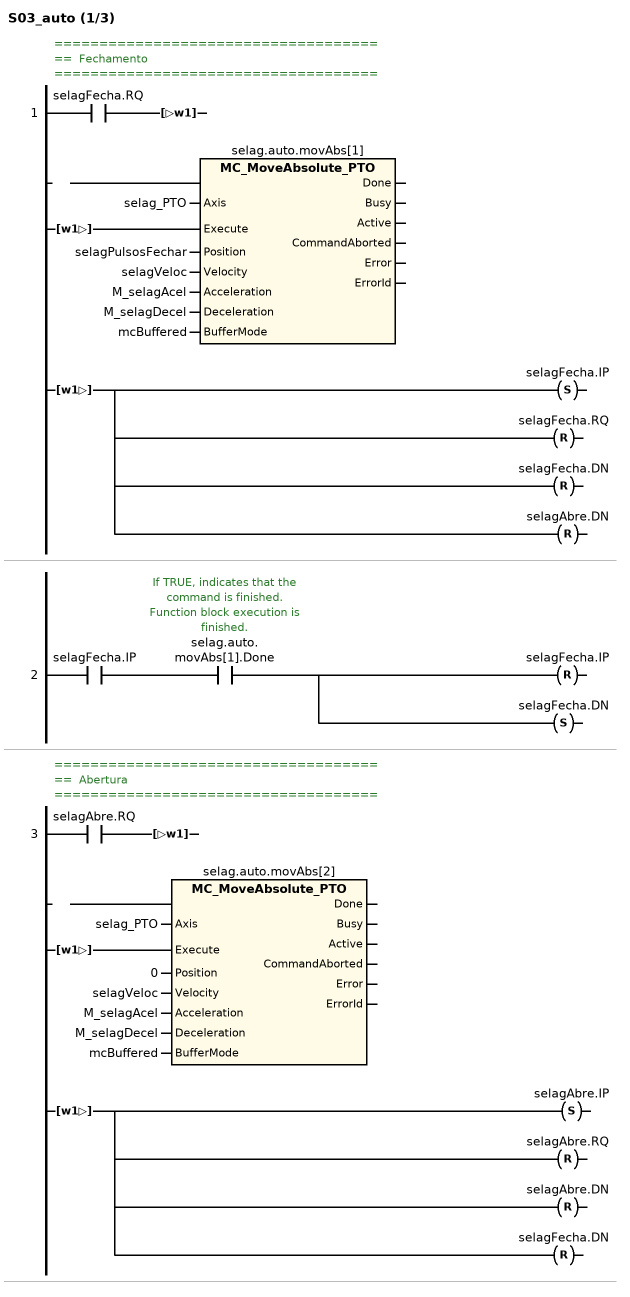
// NETWORK 1
// ====================================
// ==  Fechamento
// ====================================
_w1 := selagFecha.RQ;
selag.auto.movAbs[1](
    Axis := selag_PTO,
    Execute := _w1,
    Position := selagPulsosFechar,
    Velocity := selagVeloc,
    Acceleration := M_selagAcel,
    Deceleration := M_selagDecel,
    BufferMode := mcBuffered); // MC_MoveAbsolute_PTO
selagFecha.IP S= _w1;
selagFecha.RQ R= _w1;
selagFecha.DN R= _w1;
selagAbre.DN R= _w1;

// NETWORK 2
//   selag.auto.movAbs[1].Done: If TRUE, indicates that the command is finished. Function block execution is finished.
_w2 := selagFecha.IP AND selag.auto.movAbs[1].Done;
selagFecha.IP R= _w2;
selagFecha.DN S= _w2;

// NETWORK 3
// ====================================
// ==  Abertura
// ====================================
_w3 := selagAbre.RQ;
selag.auto.movAbs[2](
    Axis := selag_PTO,
    Execute := _w3,
    Position := 0,
    Velocity := selagVeloc,
    Acceleration := M_selagAcel,
    Deceleration := M_selagDecel,
    BufferMode := mcBuffered); // MC_MoveAbsolute_PTO
selagAbre.IP S= _w3;
selagAbre.RQ R= _w3;
selagAbre.DN R= _w3;
selagFecha.DN R= _w3;

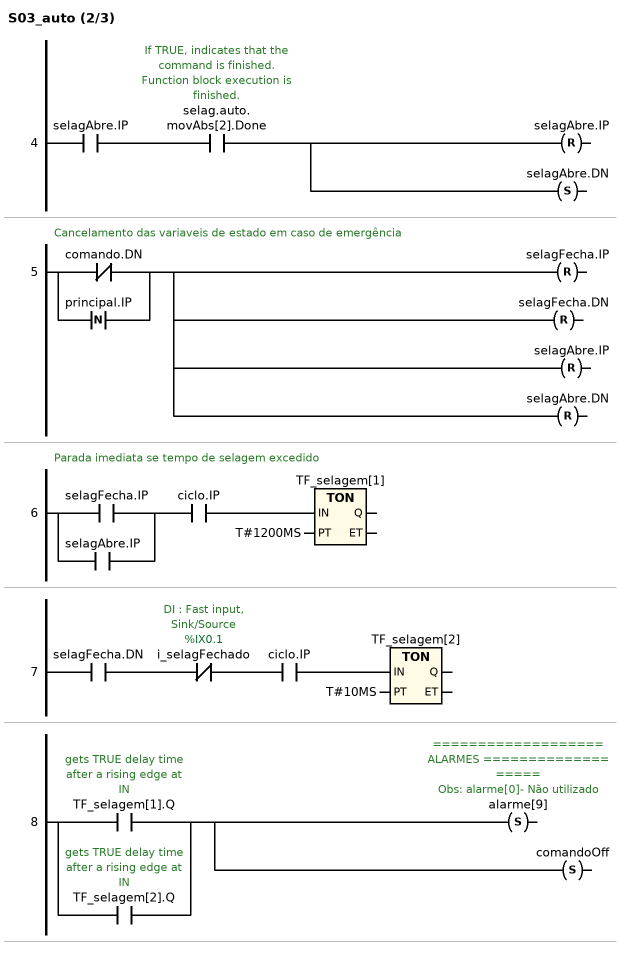
// NETWORK 4
//   selag.auto.movAbs[2].Done: If TRUE, indicates that the command is finished. Function block execution is finished.
_w4 := selagAbre.IP AND selag.auto.movAbs[2].Done;
selagAbre.IP R= _w4;
selagAbre.DN S= _w4;

// NETWORK 5
// Cancelamento das variaveis de estado em caso de emergência
_ft1(CLK := principal.IP);
_w5 := NOT comando.DN OR _ft1.Q;
selagFecha.IP R= _w5;
selagFecha.DN R= _w5;
selagAbre.IP R= _w5;
selagAbre.DN R= _w5;

// NETWORK 6
// Parada imediata se tempo de selagem excedido
TF_selagem[1](IN := (selagFecha.IP OR selagAbre.IP) AND ciclo.IP, PT := T#1200MS); // TON

// NETWORK 7
//   i_selagFechado: DI : Fast input, Sink/Source | AT %IX0.1
TF_selagem[2](IN := selagFecha.DN AND NOT i_selagFechado AND ciclo.IP, PT := T#10MS); // TON

// NETWORK 8
//   TF_selagem[1].Q: gets TRUE delay time after a rising edge at IN
//   TF_selagem[2].Q: gets TRUE delay time after a rising edge at IN
//   alarme[9]: =================== ALARMES =================== Obs: alarme[0]- Não utilizado
_w6 := TF_selagem[1].Q OR TF_selagem[2].Q;
alarme[9] S= _w6;
comandoOff S= _w6;

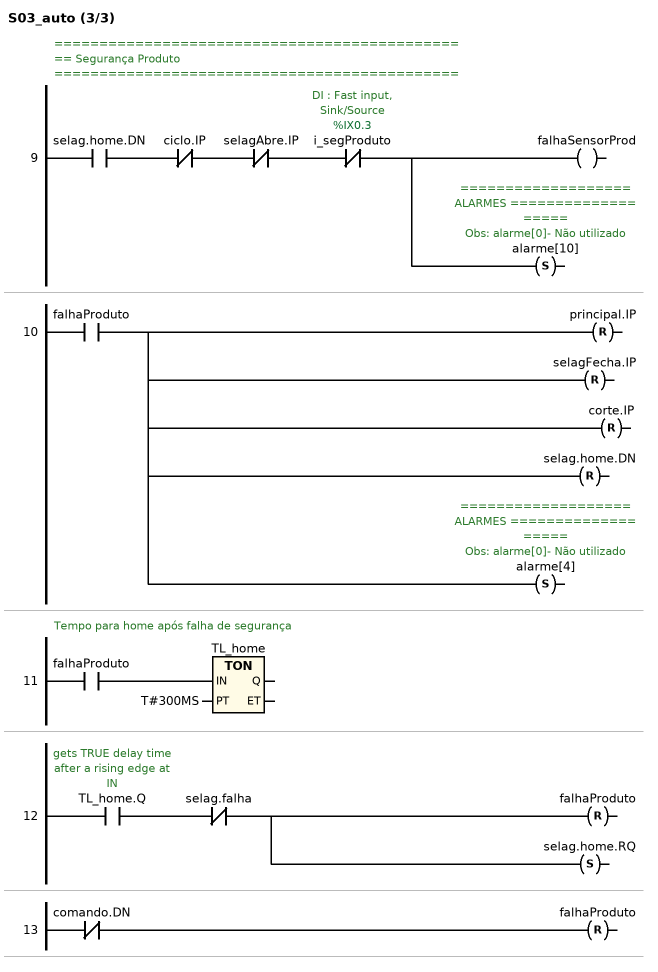
// NETWORK 9
// =============================================
// == Segurança Produto
// =============================================
//   i_segProduto: DI : Fast input, Sink/Source | AT %IX0.3
//   alarme[10]: =================== ALARMES =================== Obs: alarme[0]- Não utilizado
_w7 := selag.home.DN AND NOT ciclo.IP AND NOT selagAbre.IP AND NOT i_segProduto;
falhaSensorProd := _w7;
alarme[10] S= _w7;

// NETWORK 10
//   alarme[4]: =================== ALARMES =================== Obs: alarme[0]- Não utilizado
principal.IP R= falhaProduto;
selagFecha.IP R= falhaProduto;
corte.IP R= falhaProduto;
selag.home.DN R= falhaProduto;
alarme[4] S= falhaProduto;

// NETWORK 11
// Tempo para home após falha de segurança
TL_home(IN := falhaProduto, PT := T#300MS); // TON

// NETWORK 12
//   TL_home.Q: gets TRUE delay time after a rising edge at IN
_w8 := TL_home.Q AND NOT selag.falha;
falhaProduto R= _w8;
selag.home.RQ S= _w8;

// NETWORK 13
falhaProduto R= NOT comando.DN;

END_PROGRAM

// MyController/Application/03_Selagem/S99_calculo
PROGRAM S99_calculo
VAR
END_VAR

selag.calcula:= FALSE;

// cálculo do num pulsos/mm - 1volta motor = 47 mm
selagPulsosMm:= M_selagPulsosVolta / 47;

// cálculo das distâncias a serem percorridas
selagPulsosFechar:= REAL_TO_DINT(M_selagPosFecha * selagPulsosMm / 10);

// cálculo da velocidade
selagVeloc:= 299 * M_selagPulsosVolta * M_selagVeloc / 6000;
selagVelocHome:= 299 * M_selagPulsosVolta * M_selagVelocHome / 6000;

END_PROGRAM

// MyController/Application/04_Disco/D03_auto
PROGRAM D03_auto
VAR
	TF_foto						: TON;
END_VAR
VAR // added by the converter: edge detectors and wires of the graphical bodies
    _w1, _w2 : BOOL;
    _ft1 : F_TRIG;
END_VAR

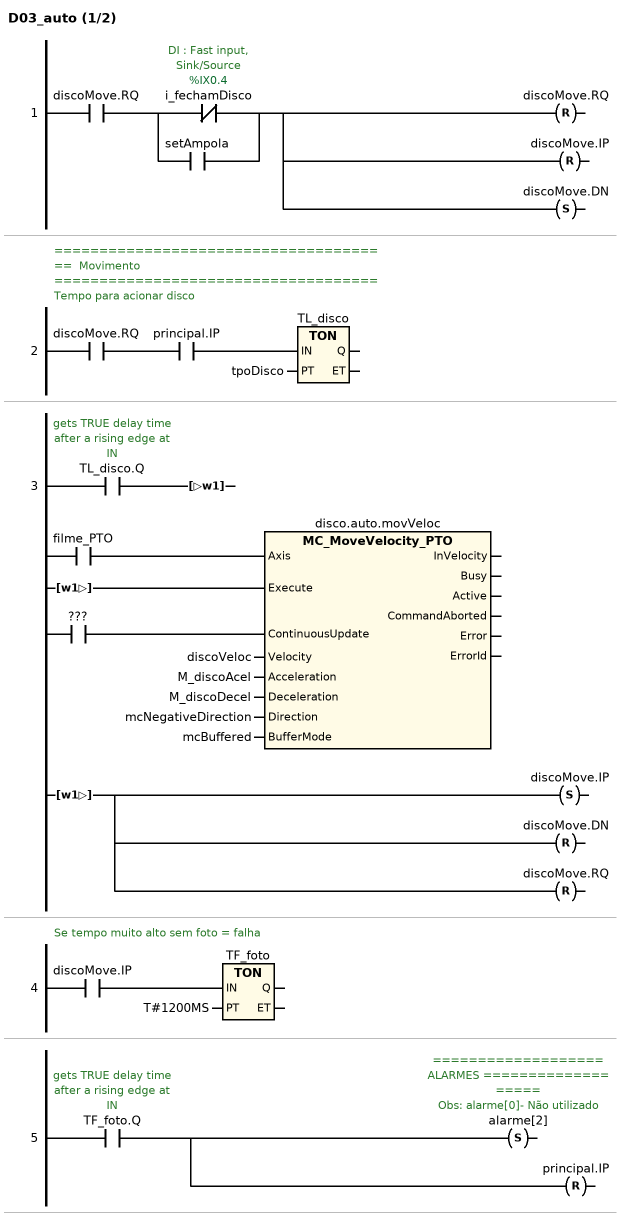
// NETWORK 1
//   i_fechamDisco: DI : Fast input, Sink/Source | AT %IX0.4
_w1 := discoMove.RQ AND (NOT i_fechamDisco OR setAmpola);
discoMove.RQ R= _w1;
discoMove.IP R= _w1;
discoMove.DN S= _w1;

// NETWORK 2
// ====================================
// ==  Movimento
// ====================================
// Tempo para acionar disco
TL_disco(IN := discoMove.RQ AND principal.IP, PT := tpoDisco); // TON

// NETWORK 3
//   TL_disco.Q: gets TRUE delay time after a rising edge at IN
disco.auto.movVeloc(
    Axis := filme_PTO,
    Execute := TL_disco.Q,
    Velocity := discoVeloc,
    Acceleration := M_discoAcel,
    Deceleration := M_discoDecel,
    Direction := mcNegativeDirection,
    BufferMode := mcBuffered); // MC_MoveVelocity_PTO
discoMove.IP S= TL_disco.Q;
discoMove.DN R= TL_disco.Q;
discoMove.RQ R= TL_disco.Q;

// NETWORK 4
// Se tempo muito alto sem foto = falha
TF_foto(IN := discoMove.IP, PT := T#1200MS); // TON

// NETWORK 5
//   TF_foto.Q: gets TRUE delay time after a rising edge at IN
//   alarme[2]: =================== ALARMES =================== Obs: alarme[0]- Não utilizado
alarme[2] S= TF_foto.Q;
principal.IP R= TF_foto.Q;

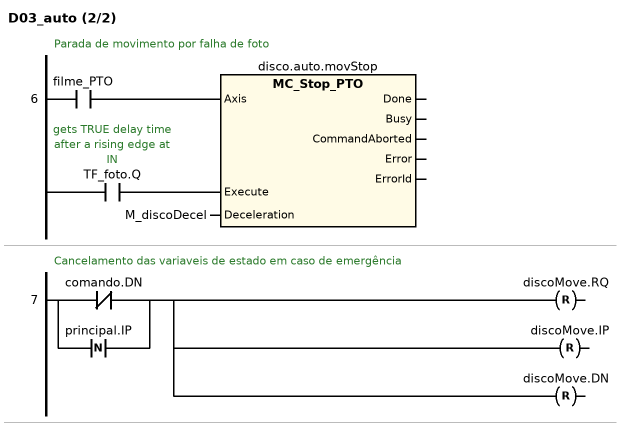
// NETWORK 6
// Parada de movimento por falha de foto
//   TF_foto.Q: gets TRUE delay time after a rising edge at IN
disco.auto.movStop(Axis := filme_PTO, Execute := TF_foto.Q, Deceleration := M_discoDecel); // MC_Stop_PTO

// NETWORK 7
// Cancelamento das variaveis de estado em caso de emergência
_ft1(CLK := principal.IP);
_w2 := NOT comando.DN OR _ft1.Q;
discoMove.RQ R= _w2;
discoMove.IP R= _w2;
discoMove.DN R= _w2;

END_PROGRAM

// MyController/Application/04_Disco/D99_calculo
PROGRAM D99_calculo
VAR
END_VAR

disco.calcula:= FALSE;

// cálculo do num pulsos/mm
discoPulsosMm:= M_discoPulsosVolta / (pi * M_diamDisco);

// cálculo das distâncias a serem percorridas
discoPulsosAposFoto:= -1 * REAL_TO_DINT(Rc[numReceita].discoMmAposFoto * discoPulsosMm);

// cálculo da velocidade
discoVeloc:= 350 * M_discoPulsosVolta * M_discoVeloc / 6000;

END_PROGRAM

// MyController/Application/05_IHM/I01_geral
PROGRAM I01_geral
VAR
	auxBit				: BOOL;
END_VAR
VAR // added by the converter: edge detectors and wires of the graphical bodies
    _rt1, _rt2, _rt3 : R_TRIG;
    _w1, _w2, _w3, _w4, _w5 : BOOL;
END_VAR

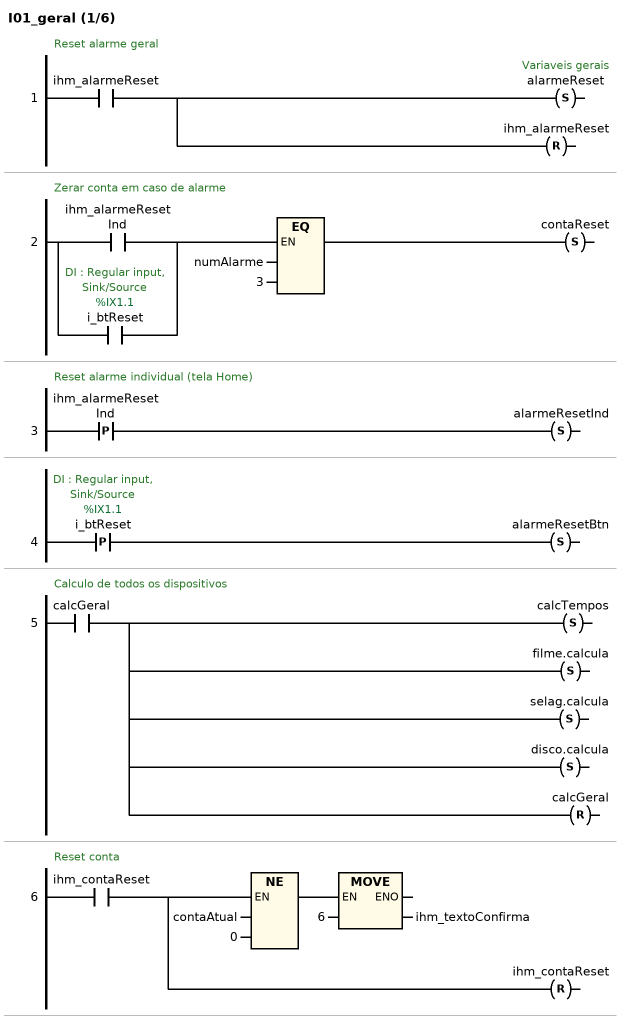
// NETWORK 1
// Reset alarme geral
//   alarmeReset: Variaveis gerais
alarmeReset S= ihm_alarmeReset;
ihm_alarmeReset R= ihm_alarmeReset;

// NETWORK 2
// Zerar conta em caso de alarme
//   i_btReset: DI : Regular input, Sink/Source | AT %IX1.1
contaReset S= (ihm_alarmeResetInd OR i_btReset) AND numAlarme = 3;

// NETWORK 3
// Reset alarme individual (tela Home)
_rt1(CLK := ihm_alarmeResetInd);
alarmeResetInd S= _rt1.Q;

// NETWORK 4
//   i_btReset: DI : Regular input, Sink/Source | AT %IX1.1
_rt2(CLK := i_btReset);
alarmeResetBtn S= _rt2.Q;

// NETWORK 5
// Calculo de todos os dispositivos
calcTempos S= calcGeral;
filme.calcula S= calcGeral;
selag.calcula S= calcGeral;
disco.calcula S= calcGeral;
calcGeral R= calcGeral;

// NETWORK 6
// Reset conta
_w1 := ihm_contaReset;
IF _w1 AND contaAtual <> 0 THEN ihm_textoConfirma := 6; END_IF
ihm_contaReset R= _w1;

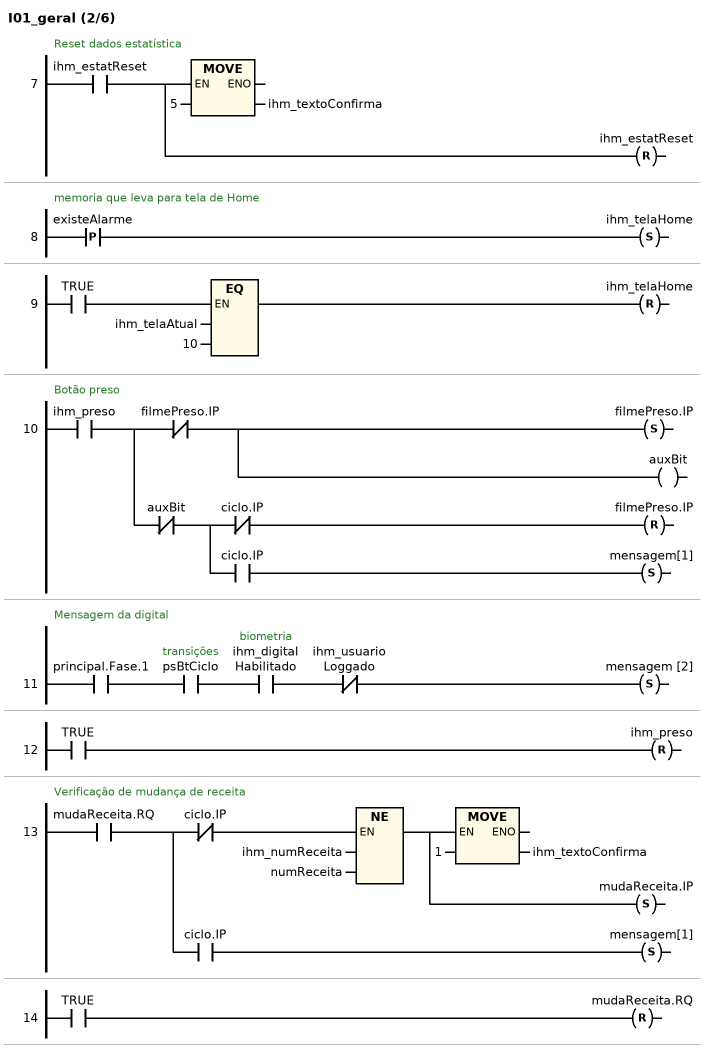
// NETWORK 7
// Reset dados estatística
_w2 := ihm_estatReset;
IF _w2 THEN ihm_textoConfirma := 5; END_IF
ihm_estatReset R= _w2;

// NETWORK 8
// memoria que leva para tela de Home
_rt3(CLK := existeAlarme);
ihm_telaHome S= _rt3.Q;

// NETWORK 9
ihm_telaHome R= ihm_telaAtual = 10;

// NETWORK 10
// Botão preso
_w3 := ihm_preso AND NOT filmePreso.IP;
filmePreso.IP S= _w3;
auxBit := _w3;
_w4 := ihm_preso AND NOT auxBit;
filmePreso.IP R= _w4 AND NOT ciclo.IP;
mensagem[1] S= _w4 AND ciclo.IP;

// NETWORK 11
//  Mensagem da digital
//   psBtCiclo: transições
//   ihm_digitalHabilitado: biometria
mensagem [2] S= principal.Fase.1 AND psBtCiclo AND ihm_digitalHabilitado AND NOT ihm_usuarioLoggado;

// NETWORK 12
ihm_preso R= TRUE;

// NETWORK 13
// Verificação de mudança de receita
_w5 := mudaReceita.RQ AND NOT ciclo.IP AND ihm_numReceita <> numReceita;
IF _w5 THEN ihm_textoConfirma := 1; END_IF
mudaReceita.IP S= _w5;
mensagem[1] S= mudaReceita.RQ AND ciclo.IP;

// NETWORK 14
mudaReceita.RQ R= TRUE;

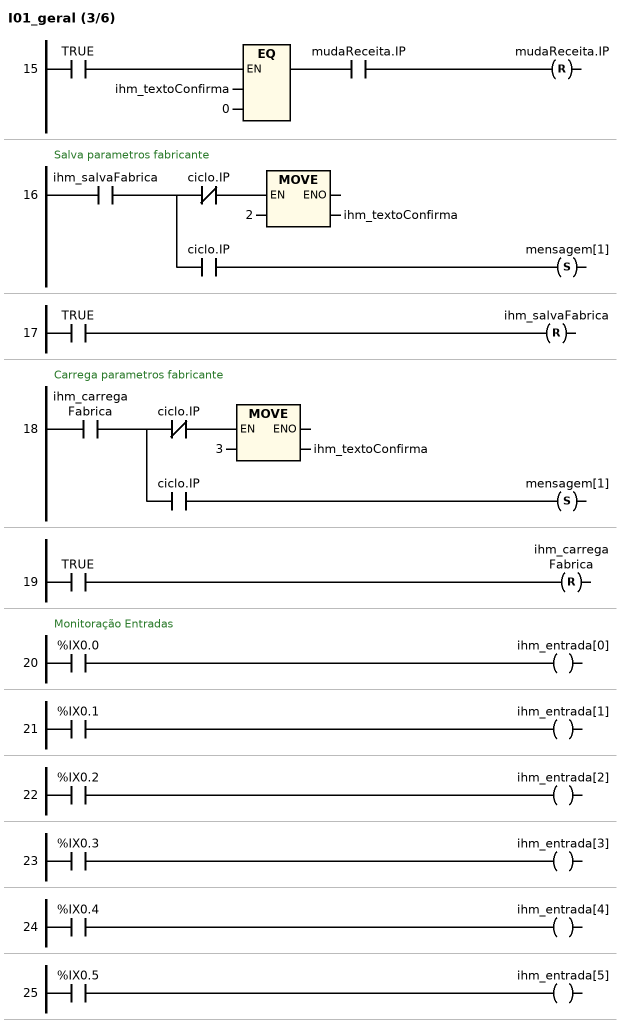
// NETWORK 15
mudaReceita.IP R= ihm_textoConfirma = 0 AND mudaReceita.IP;

// NETWORK 16
// Salva parametros fabricante
IF ihm_salvaFabrica AND NOT ciclo.IP THEN ihm_textoConfirma := 2; END_IF
mensagem[1] S= ihm_salvaFabrica AND ciclo.IP;

// NETWORK 17
ihm_salvaFabrica R= TRUE;

// NETWORK 18
// Carrega parametros fabricante
IF ihm_carregaFabrica AND NOT ciclo.IP THEN ihm_textoConfirma := 3; END_IF
mensagem[1] S= ihm_carregaFabrica AND ciclo.IP;

// NETWORK 19
ihm_carregaFabrica R= TRUE;

// NETWORK 20
// Monitoração Entradas
ihm_entrada[0] := %IX0.0;

// NETWORK 21
ihm_entrada[1] := %IX0.1;

// NETWORK 22
ihm_entrada[2] := %IX0.2;

// NETWORK 23
ihm_entrada[3] := %IX0.3;

// NETWORK 24
ihm_entrada[4] := %IX0.4;

// NETWORK 25
ihm_entrada[5] := %IX0.5;

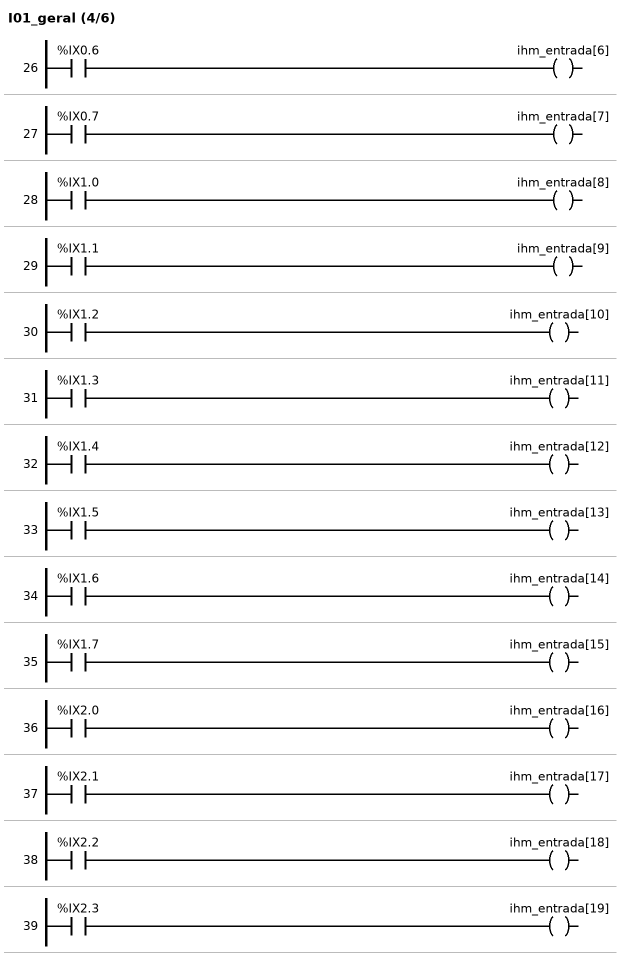
// NETWORK 26
ihm_entrada[6] := %IX0.6;

// NETWORK 27
ihm_entrada[7] := %IX0.7;

// NETWORK 28
ihm_entrada[8] := %IX1.0;

// NETWORK 29
ihm_entrada[9] := %IX1.1;

// NETWORK 30
ihm_entrada[10] := %IX1.2;

// NETWORK 31
ihm_entrada[11] := %IX1.3;

// NETWORK 32
ihm_entrada[12] := %IX1.4;

// NETWORK 33
ihm_entrada[13] := %IX1.5;

// NETWORK 34
ihm_entrada[14] := %IX1.6;

// NETWORK 35
ihm_entrada[15] := %IX1.7;

// NETWORK 36
ihm_entrada[16] := %IX2.0;

// NETWORK 37
ihm_entrada[17] := %IX2.1;

// NETWORK 38
ihm_entrada[18] := %IX2.2;

// NETWORK 39
ihm_entrada[19] := %IX2.3;

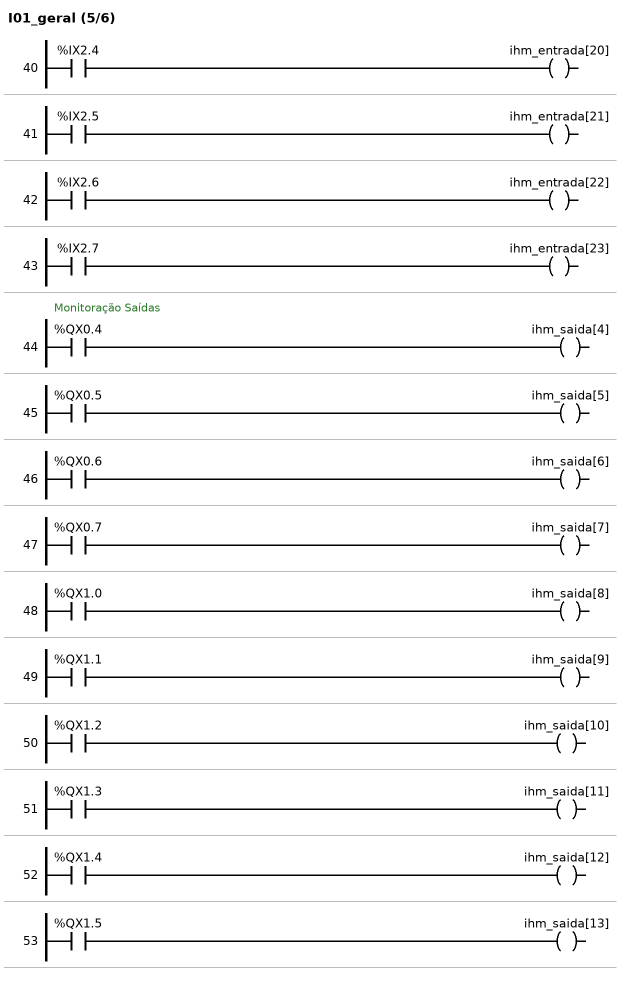
// NETWORK 40
ihm_entrada[20] := %IX2.4;

// NETWORK 41
ihm_entrada[21] := %IX2.5;

// NETWORK 42
ihm_entrada[22] := %IX2.6;

// NETWORK 43
ihm_entrada[23] := %IX2.7;

// NETWORK 44
// Monitoração Saídas
ihm_saida[4] := %QX0.4;

// NETWORK 45
ihm_saida[5] := %QX0.5;

// NETWORK 46
ihm_saida[6] := %QX0.6;

// NETWORK 47
ihm_saida[7] := %QX0.7;

// NETWORK 48
ihm_saida[8] := %QX1.0;

// NETWORK 49
ihm_saida[9] := %QX1.1;

// NETWORK 50
ihm_saida[10] := %QX1.2;

// NETWORK 51
ihm_saida[11] := %QX1.3;

// NETWORK 52
ihm_saida[12] := %QX1.4;

// NETWORK 53
ihm_saida[13] := %QX1.5;

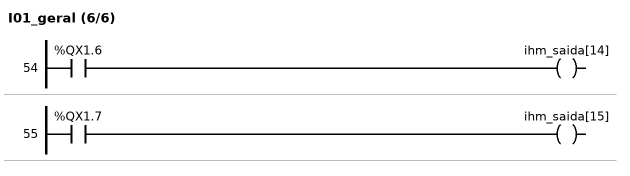
// NETWORK 54
ihm_saida[14] := %QX1.6;

// NETWORK 55
ihm_saida[15] := %QX1.7;

END_PROGRAM

// MyController/Application/05_IHM/I02_alarmes
PROGRAM I02_alarmes
VAR
	auxExisteAlarme					: BOOL;
	delayAlarme						: TON;
	memAlarme						: ARRAY[0..99] OF BOOL;
	p0								: SINT;
END_VAR


CASE alarmes.Fase OF
(*====================================
  ==  Fase 0 - alarmes 1 a 50 (0 não existe)
  ====================================*)
0:
	auxExisteAlarme:= FALSE;
	FOR p0:= 1 TO 50 DO
		IF alarme[p0] THEN
			memAlarme[p0]:= TRUE;
			auxExisteAlarme:= TRUE;
			
			IF numAlarme = 0 THEN
				numAlarme:= p0;				// pega o numero do primeiro alarme que ocorre
			END_IF
		END_IF
		
		IF numAlarme = p0 THEN
			IF alarme[p0] = 0 THEN			// verifica se o alarme que ocorreu continua ativo
				numAlarme:= 0;
			END_IF
		END_IF
	END_FOR
	alarmes.Fase:= 10;

	
(*====================================
  ==  Fase 10 - passa alarmes para ihm	
  ====================================*)
10:
	FOR p0:= 1 TO 50 DO
		ihm_alarme[p0]:= memAlarme[p0];
		memAlarme[p0]:= FALSE;
	END_FOR
	alarmes.Fase:= 11;
	
	
(*====================================
  ==  Fase 11 - verifica cancela alarmes pela IHM
  ====================================*)	
11:
	existeAlarme:= auxExisteAlarme;
	IF alarmeReset THEN
		alarmes.Fase:= 12;
	ELSE
		IF alarmeResetInd OR (alarmeResetBtn AND comando.DN) THEN
			alarme[numAlarme]:= FALSE;
			alarmeResetInd:= FALSE;
			alarmeResetBtn:= FALSE;
		END_IF
		alarmes.Fase:= 0;
	END_IF

	
(*====================================
  ==  Fase 12 - cancela alarmes	
  ====================================*)
12:
	alarmeReset:= FALSE;
	FOR p0:= 1 TO 50 DO
		alarme[p0]:= 0;
	END_FOR
	alarmes.Fase:= 13;
	

(*====================================
  ==  Fase 13 - espera 100ms para atualização dos bits de alarmes pelo controle
  ====================================*)	
13:
	IF delayAlarme.Q THEN
		alarmes.Fase:= 0;
	END_IF
	delayAlarme(IN:= alarmes.Fase= 13, PT:= T#100MS);

END_CASE

END_PROGRAM

// MyController/Application/05_IHM/I03_mensagens
PROGRAM I03_mensagens
VAR
	delayMensag						: TON;
	mensagens						: _exec_bits;
	p1								: DINT;
END_VAR


IF NOT mensagens.RQ THEN
	FOR p1:= 1 TO 50 DO
		IF mensagem[p1] = TRUE THEN
			mensagem[p1]:= 0;
			ihm_mensagem:= p1;
			mensagens.RQ:= TRUE;
		END_IF
	END_FOR
END_IF


// Tempo de cada mensagem na tela
delayMensag(IN := ihm_bannerMensagem, PT:= T#2500MS);
IF delayMensag.Q THEN
	mensagens.RQ:= FALSE;
	ihm_mensagem:= 0;
END_IF


ihm_bannerMensagem:= mensagens.RQ AND NOT ihm_bannerConfirma;

END_PROGRAM

// MyController/Application/05_IHM/I06_textoConfirma
PROGRAM I06_textoConfirma
VAR
END_VAR
VAR // added by the converter: edge detectors and wires of the graphical bodies
    _w1, _w2, _w3 : BOOL;
END_VAR
